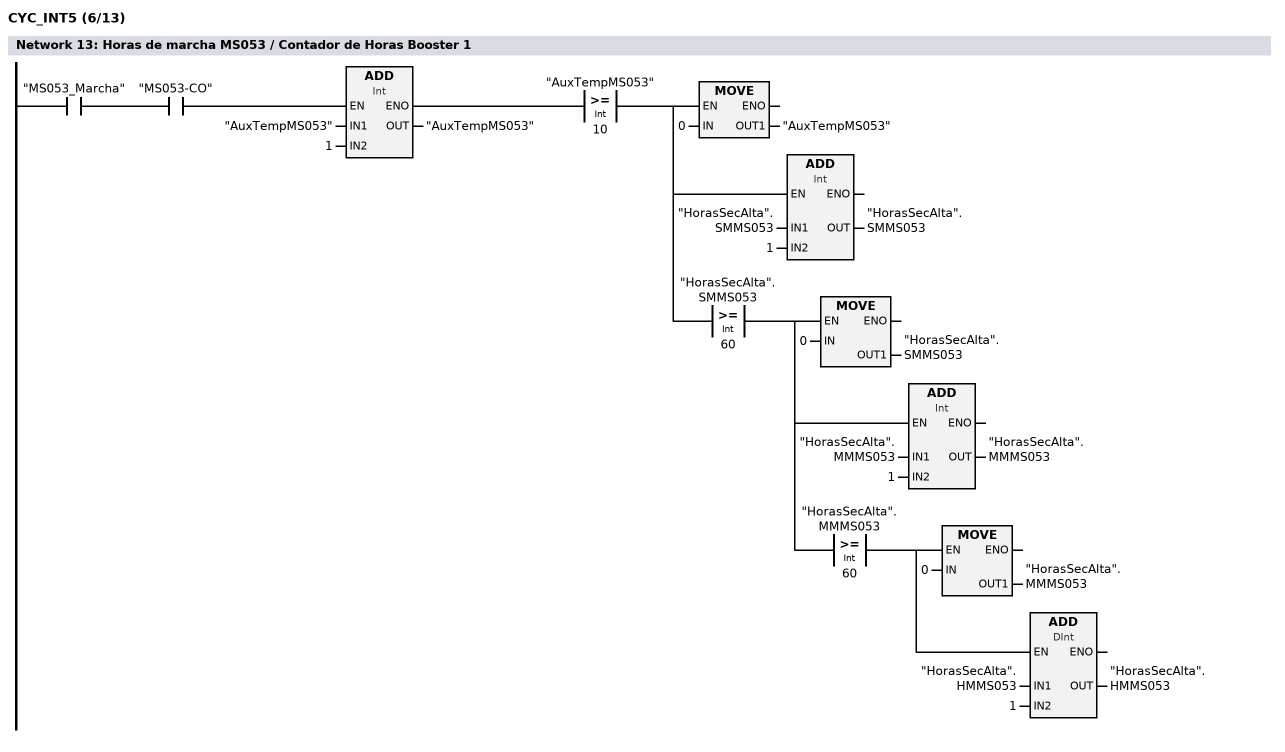
   RUNG wire#powerrail
      Contact( "MS053_Marcha" )
      Contact( "MS053-CO" )
      { S7_Templates := "SrcType := Int"; S7_GenerateENO := "TRUE" } Add(in1 := "AuxTempMS053", in2 := 1, out => "AuxTempMS053")
      { S7_Templates := "SrcType := Int" } GE_Contact(in1 := "AuxTempMS053", in2 := 10)
      wire#w1
      { S7_GenerateENO := "TRUE" } Move(in := 0, out1 => "AuxTempMS053")
   END_RUNG
   RUNG wire#w1
      { S7_Templates := "SrcType := Int"; S7_GenerateENO := "TRUE" } Add(in1 := "HorasSecAlta".SMMS053, in2 := 1, out => "HorasSecAlta".SMMS053)
   END_RUNG
   RUNG wire#w1
      { S7_Templates := "SrcType := Int" } GE_Contact(in1 := "HorasSecAlta".SMMS053, in2 := 60)
      wire#w2
      { S7_GenerateENO := "TRUE" } Move(in := 0, out1 => "HorasSecAlta".SMMS053)
   END_RUNG
   RUNG wire#w2
      { S7_Templates := "SrcType := Int"; S7_GenerateENO := "TRUE" } Add(in1 := "HorasSecAlta".MMMS053, in2 := 1, out => "HorasSecAlta".MMMS053)
   END_RUNG
   RUNG wire#w2
      { S7_Templates := "SrcType := Int" } GE_Contact(in1 := "HorasSecAlta".MMMS053, in2 := 60)
      wire#w3
      { S7_GenerateENO := "TRUE" } Move(in := 0, out1 => "HorasSecAlta".MMMS053)
   END_RUNG
   RUNG wire#w3
      { S7_Templates := "SrcType := DInt"; S7_GenerateENO := "TRUE" } Add(in1 := "HorasSecAlta".HMMS053, in2 := 1, out => "HorasSecAlta".HMMS053)
   END_RUNG
   // the same network as SCL:
   // ENO of a box is taken as its EN; it also drops when the box reports an error
   #_w1 := "MS053_Marcha" AND "MS053-CO";
   IF #_w1 THEN "AuxTempMS053" := "AuxTempMS053" + 1; END_IF;
   #_w2 := #_w1 AND ("AuxTempMS053" >= 10);
   IF #_w2 THEN
       "AuxTempMS053" := 0;
       "HorasSecAlta".SMMS053 := "HorasSecAlta".SMMS053 + 1;
   END_IF;
   #_w3 := #_w2 AND ("HorasSecAlta".SMMS053 >= 60);
   IF #_w3 THEN
       "HorasSecAlta".SMMS053 := 0;
       "HorasSecAlta".MMMS053 := "HorasSecAlta".MMMS053 + 1;
   END_IF;
   #_w4 := #_w3 AND ("HorasSecAlta".MMMS053 >= 60);
   IF #_w4 THEN
       "HorasSecAlta".MMMS053 := 0;
       "HorasSecAlta".HMMS053 := "HorasSecAlta".HMMS053 + 1;
   END_IF;
END_REGION

REGION Network 14: Horas de marcha MS054 / Contador de Horas Booster 1
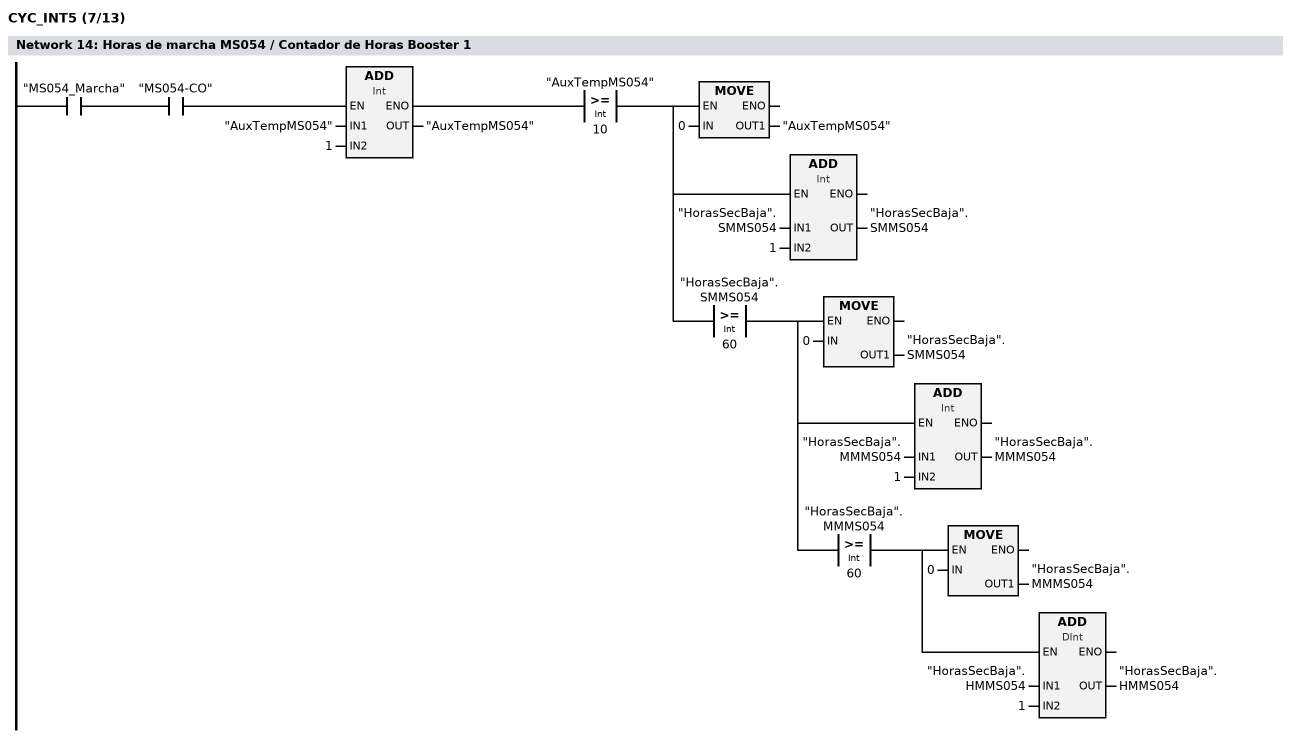
   RUNG wire#powerrail
      Contact( "MS054_Marcha" )
      Contact( "MS054-CO" )
      { S7_Templates := "SrcType := Int"; S7_GenerateENO := "TRUE" } Add(in1 := "AuxTempMS054", in2 := 1, out => "AuxTempMS054")
      { S7_Templates := "SrcType := Int" } GE_Contact(in1 := "AuxTempMS054", in2 := 10)
      wire#w1
      { S7_GenerateENO := "TRUE" } Move(in := 0, out1 => "AuxTempMS054")
   END_RUNG
   RUNG wire#w1
      { S7_Templates := "SrcType := Int"; S7_GenerateENO := "TRUE" } Add(in1 := "HorasSecBaja".SMMS054, in2 := 1, out => "HorasSecBaja".SMMS054)
   END_RUNG
   RUNG wire#w1
      { S7_Templates := "SrcType := Int" } GE_Contact(in1 := "HorasSecBaja".SMMS054, in2 := 60)
      wire#w2
      { S7_GenerateENO := "TRUE" } Move(in := 0, out1 => "HorasSecBaja".SMMS054)
   END_RUNG
   RUNG wire#w2
      { S7_Templates := "SrcType := Int"; S7_GenerateENO := "TRUE" } Add(in1 := "HorasSecBaja".MMMS054, in2 := 1, out => "HorasSecBaja".MMMS054)
   END_RUNG
   RUNG wire#w2
      { S7_Templates := "SrcType := Int" } GE_Contact(in1 := "HorasSecBaja".MMMS054, in2 := 60)
      wire#w3
      { S7_GenerateENO := "TRUE" } Move(in := 0, out1 => "HorasSecBaja".MMMS054)
   END_RUNG
   RUNG wire#w3
      { S7_Templates := "SrcType := DInt"; S7_GenerateENO := "TRUE" } Add(in1 := "HorasSecBaja".HMMS054, in2 := 1, out => "HorasSecBaja".HMMS054)
   END_RUNG
   // the same network as SCL:
   // ENO of a box is taken as its EN; it also drops when the box reports an error
   #_w1 := "MS054_Marcha" AND "MS054-CO";
   IF #_w1 THEN "AuxTempMS054" := "AuxTempMS054" + 1; END_IF;
   #_w2 := #_w1 AND ("AuxTempMS054" >= 10);
   IF #_w2 THEN
       "AuxTempMS054" := 0;
       "HorasSecBaja".SMMS054 := "HorasSecBaja".SMMS054 + 1;
   END_IF;
   #_w3 := #_w2 AND ("HorasSecBaja".SMMS054 >= 60);
   IF #_w3 THEN
       "HorasSecBaja".SMMS054 := 0;
       "HorasSecBaja".MMMS054 := "HorasSecBaja".MMMS054 + 1;
   END_IF;
   #_w4 := #_w3 AND ("HorasSecBaja".MMMS054 >= 60);
   IF #_w4 THEN
       "HorasSecBaja".MMMS054 := 0;
       "HorasSecBaja".HMMS054 := "HorasSecBaja".HMMS054 + 1;
   END_IF;
END_REGION

REGION Network 15: Horas de marcha MS055 / Contador de Horas Booster 1
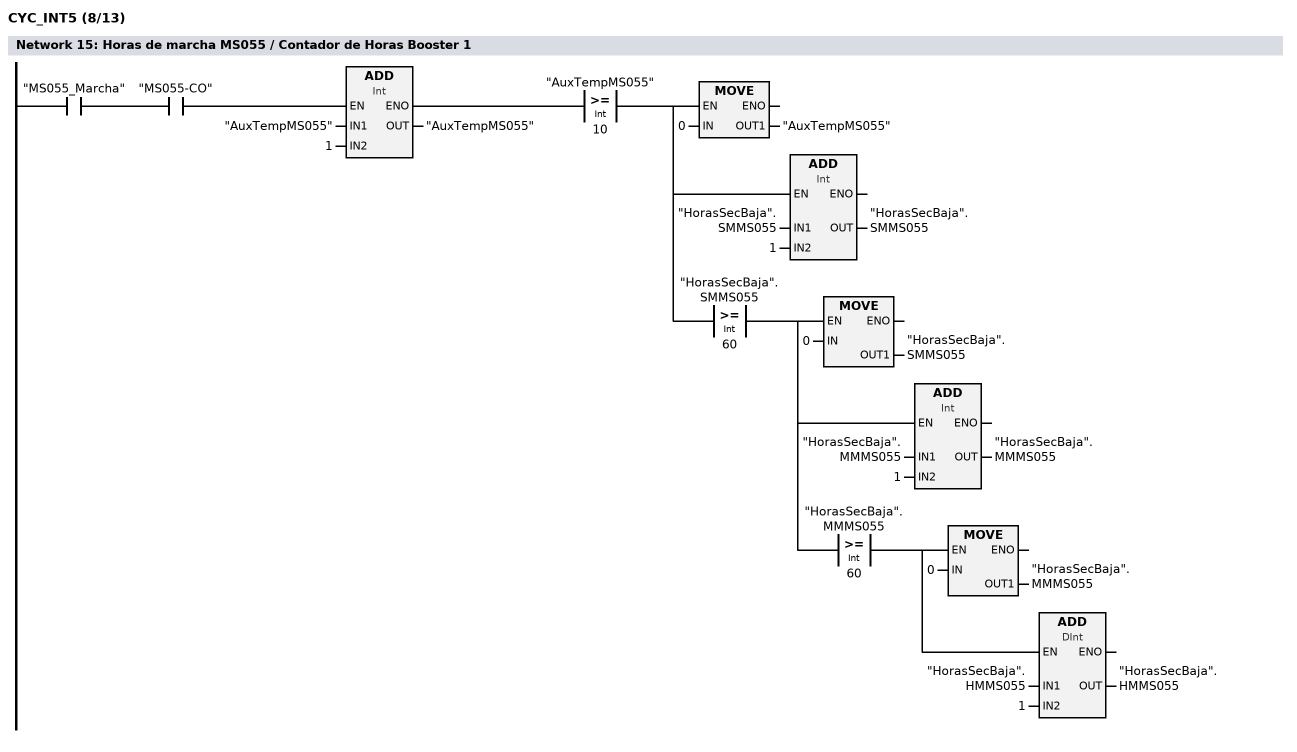
   RUNG wire#powerrail
      Contact( "MS055_Marcha" )
      Contact( "MS055-CO" )
      { S7_Templates := "SrcType := Int"; S7_GenerateENO := "TRUE" } Add(in1 := "AuxTempMS055", in2 := 1, out => "AuxTempMS055")
      { S7_Templates := "SrcType := Int" } GE_Contact(in1 := "AuxTempMS055", in2 := 10)
      wire#w1
      { S7_GenerateENO := "TRUE" } Move(in := 0, out1 => "AuxTempMS055")
   END_RUNG
   RUNG wire#w1
      { S7_Templates := "SrcType := Int"; S7_GenerateENO := "TRUE" } Add(in1 := "HorasSecBaja".SMMS055, in2 := 1, out => "HorasSecBaja".SMMS055)
   END_RUNG
   RUNG wire#w1
      { S7_Templates := "SrcType := Int" } GE_Contact(in1 := "HorasSecBaja".SMMS055, in2 := 60)
      wire#w2
      { S7_GenerateENO := "TRUE" } Move(in := 0, out1 => "HorasSecBaja".SMMS055)
   END_RUNG
   RUNG wire#w2
      { S7_Templates := "SrcType := Int"; S7_GenerateENO := "TRUE" } Add(in1 := "HorasSecBaja".MMMS055, in2 := 1, out => "HorasSecBaja".MMMS055)
   END_RUNG
   RUNG wire#w2
      { S7_Templates := "SrcType := Int" } GE_Contact(in1 := "HorasSecBaja".MMMS055, in2 := 60)
      wire#w3
      { S7_GenerateENO := "TRUE" } Move(in := 0, out1 => "HorasSecBaja".MMMS055)
   END_RUNG
   RUNG wire#w3
      { S7_Templates := "SrcType := DInt"; S7_GenerateENO := "TRUE" } Add(in1 := "HorasSecBaja".HMMS055, in2 := 1, out => "HorasSecBaja".HMMS055)
   END_RUNG
   // the same network as SCL:
   // ENO of a box is taken as its EN; it also drops when the box reports an error
   #_w1 := "MS055_Marcha" AND "MS055-CO";
   IF #_w1 THEN "AuxTempMS055" := "AuxTempMS055" + 1; END_IF;
   #_w2 := #_w1 AND ("AuxTempMS055" >= 10);
   IF #_w2 THEN
       "AuxTempMS055" := 0;
       "HorasSecBaja".SMMS055 := "HorasSecBaja".SMMS055 + 1;
   END_IF;
   #_w3 := #_w2 AND ("HorasSecBaja".SMMS055 >= 60);
   IF #_w3 THEN
       "HorasSecBaja".SMMS055 := 0;
       "HorasSecBaja".MMMS055 := "HorasSecBaja".MMMS055 + 1;
   END_IF;
   #_w4 := #_w3 AND ("HorasSecBaja".MMMS055 >= 60);
   IF #_w4 THEN
       "HorasSecBaja".MMMS055 := 0;
       "HorasSecBaja".HMMS055 := "HorasSecBaja".HMMS055 + 1;
   END_IF;
END_REGION

REGION Network 16: Horas de marcha MC060 / Contador de Horas Booster 1
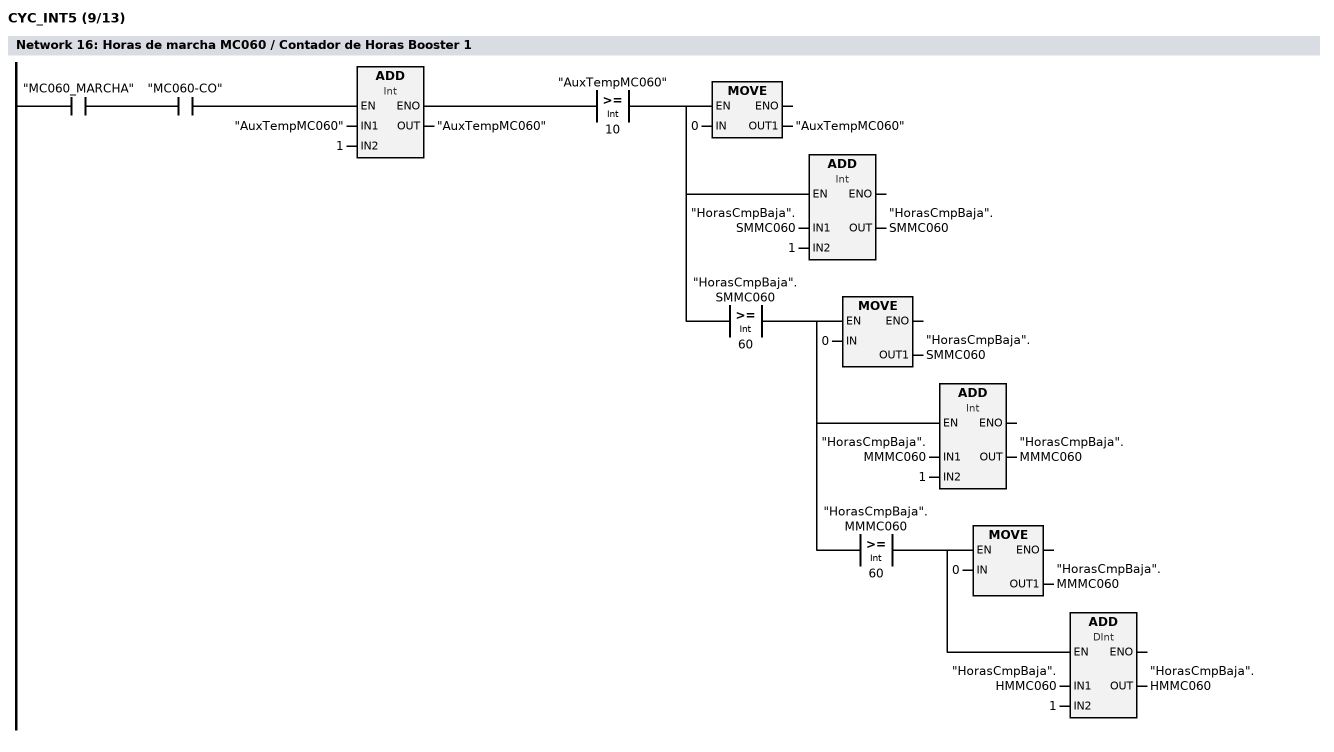
   RUNG wire#powerrail
      Contact( "MC060_MARCHA" )
      Contact( "MC060-CO" )
      { S7_Templates := "SrcType := Int"; S7_GenerateENO := "TRUE" } Add(in1 := "AuxTempMC060", in2 := 1, out => "AuxTempMC060")
      { S7_Templates := "SrcType := Int" } GE_Contact(in1 := "AuxTempMC060", in2 := 10)
      wire#w1
      { S7_GenerateENO := "TRUE" } Move(in := 0, out1 => "AuxTempMC060")
   END_RUNG
   RUNG wire#w1
      { S7_Templates := "SrcType := Int"; S7_GenerateENO := "TRUE" } Add(in1 := "HorasCmpBaja".SMMC060, in2 := 1, out => "HorasCmpBaja".SMMC060)
   END_RUNG
   RUNG wire#w1
      { S7_Templates := "SrcType := Int" } GE_Contact(in1 := "HorasCmpBaja".SMMC060, in2 := 60)
      wire#w2
      { S7_GenerateENO := "TRUE" } Move(in := 0, out1 => "HorasCmpBaja".SMMC060)
   END_RUNG
   RUNG wire#w2
      { S7_Templates := "SrcType := Int"; S7_GenerateENO := "TRUE" } Add(in1 := "HorasCmpBaja".MMMC060, in2 := 1, out => "HorasCmpBaja".MMMC060)
   END_RUNG
   RUNG wire#w2
      { S7_Templates := "SrcType := Int" } GE_Contact(in1 := "HorasCmpBaja".MMMC060, in2 := 60)
      wire#w3
      { S7_GenerateENO := "TRUE" } Move(in := 0, out1 => "HorasCmpBaja".MMMC060)
   END_RUNG
   RUNG wire#w3
      { S7_Templates := "SrcType := DInt"; S7_GenerateENO := "TRUE" } Add(in1 := "HorasCmpBaja".HMMC060, in2 := 1, out => "HorasCmpBaja".HMMC060)
   END_RUNG
   // the same network as SCL:
   // ENO of a box is taken as its EN; it also drops when the box reports an error
   #_w1 := "MC060_MARCHA" AND "MC060-CO";
   IF #_w1 THEN "AuxTempMC060" := "AuxTempMC060" + 1; END_IF;
   #_w2 := #_w1 AND ("AuxTempMC060" >= 10);
   IF #_w2 THEN
       "AuxTempMC060" := 0;
       "HorasCmpBaja".SMMC060 := "HorasCmpBaja".SMMC060 + 1;
   END_IF;
   #_w3 := #_w2 AND ("HorasCmpBaja".SMMC060 >= 60);
   IF #_w3 THEN
       "HorasCmpBaja".SMMC060 := 0;
       "HorasCmpBaja".MMMC060 := "HorasCmpBaja".MMMC060 + 1;
   END_IF;
   #_w4 := #_w3 AND ("HorasCmpBaja".MMMC060 >= 60);
   IF #_w4 THEN
       "HorasCmpBaja".MMMC060 := 0;
       "HorasCmpBaja".HMMC060 := "HorasCmpBaja".HMMC060 + 1;
   END_IF;
END_REGION

REGION Network 17: Horas de marcha MC061 / Contador de Horas Booster 1
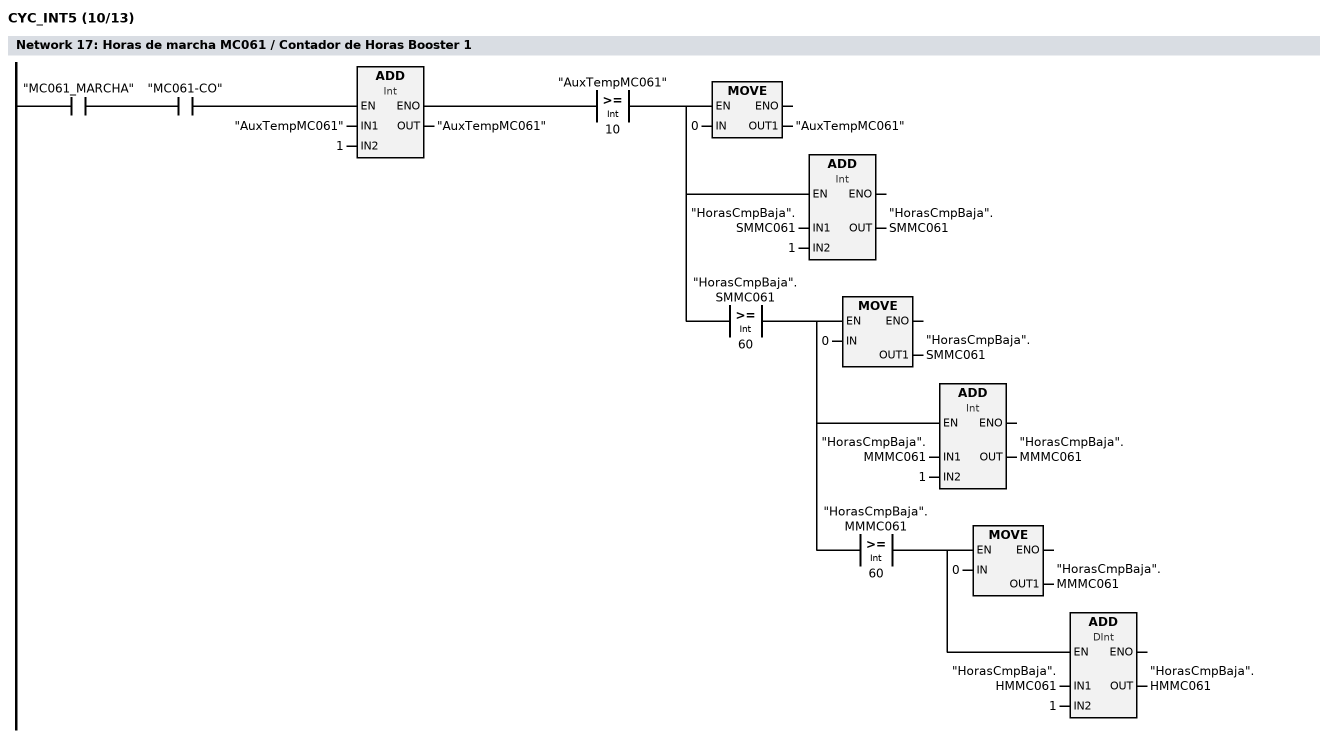
   RUNG wire#powerrail
      Contact( "MC061_MARCHA" )
      Contact( "MC061-CO" )
      { S7_Templates := "SrcType := Int"; S7_GenerateENO := "TRUE" } Add(in1 := "AuxTempMC061", in2 := 1, out => "AuxTempMC061")
      { S7_Templates := "SrcType := Int" } GE_Contact(in1 := "AuxTempMC061", in2 := 10)
      wire#w1
      { S7_GenerateENO := "TRUE" } Move(in := 0, out1 => "AuxTempMC061")
   END_RUNG
   RUNG wire#w1
      { S7_Templates := "SrcType := Int"; S7_GenerateENO := "TRUE" } Add(in1 := "HorasCmpBaja".SMMC061, in2 := 1, out => "HorasCmpBaja".SMMC061)
   END_RUNG
   RUNG wire#w1
      { S7_Templates := "SrcType := Int" } GE_Contact(in1 := "HorasCmpBaja".SMMC061, in2 := 60)
      wire#w2
      { S7_GenerateENO := "TRUE" } Move(in := 0, out1 => "HorasCmpBaja".SMMC061)
   END_RUNG
   RUNG wire#w2
      { S7_Templates := "SrcType := Int"; S7_GenerateENO := "TRUE" } Add(in1 := "HorasCmpBaja".MMMC061, in2 := 1, out => "HorasCmpBaja".MMMC061)
   END_RUNG
   RUNG wire#w2
      { S7_Templates := "SrcType := Int" } GE_Contact(in1 := "HorasCmpBaja".MMMC061, in2 := 60)
      wire#w3
      { S7_GenerateENO := "TRUE" } Move(in := 0, out1 => "HorasCmpBaja".MMMC061)
   END_RUNG
   RUNG wire#w3
      { S7_Templates := "SrcType := DInt"; S7_GenerateENO := "TRUE" } Add(in1 := "HorasCmpBaja".HMMC061, in2 := 1, out => "HorasCmpBaja".HMMC061)
   END_RUNG
   // the same network as SCL:
   // ENO of a box is taken as its EN; it also drops when the box reports an error
   #_w1 := "MC061_MARCHA" AND "MC061-CO";
   IF #_w1 THEN "AuxTempMC061" := "AuxTempMC061" + 1; END_IF;
   #_w2 := #_w1 AND ("AuxTempMC061" >= 10);
   IF #_w2 THEN
       "AuxTempMC061" := 0;
       "HorasCmpBaja".SMMC061 := "HorasCmpBaja".SMMC061 + 1;
   END_IF;
   #_w3 := #_w2 AND ("HorasCmpBaja".SMMC061 >= 60);
   IF #_w3 THEN
       "HorasCmpBaja".SMMC061 := 0;
       "HorasCmpBaja".MMMC061 := "HorasCmpBaja".MMMC061 + 1;
   END_IF;
   #_w4 := #_w3 AND ("HorasCmpBaja".MMMC061 >= 60);
   IF #_w4 THEN
       "HorasCmpBaja".MMMC061 := 0;
       "HorasCmpBaja".HMMC061 := "HorasCmpBaja".HMMC061 + 1;
   END_IF;
END_REGION

REGION Network 18: Horas de marcha MC062 / Contador de Horas Booster 1
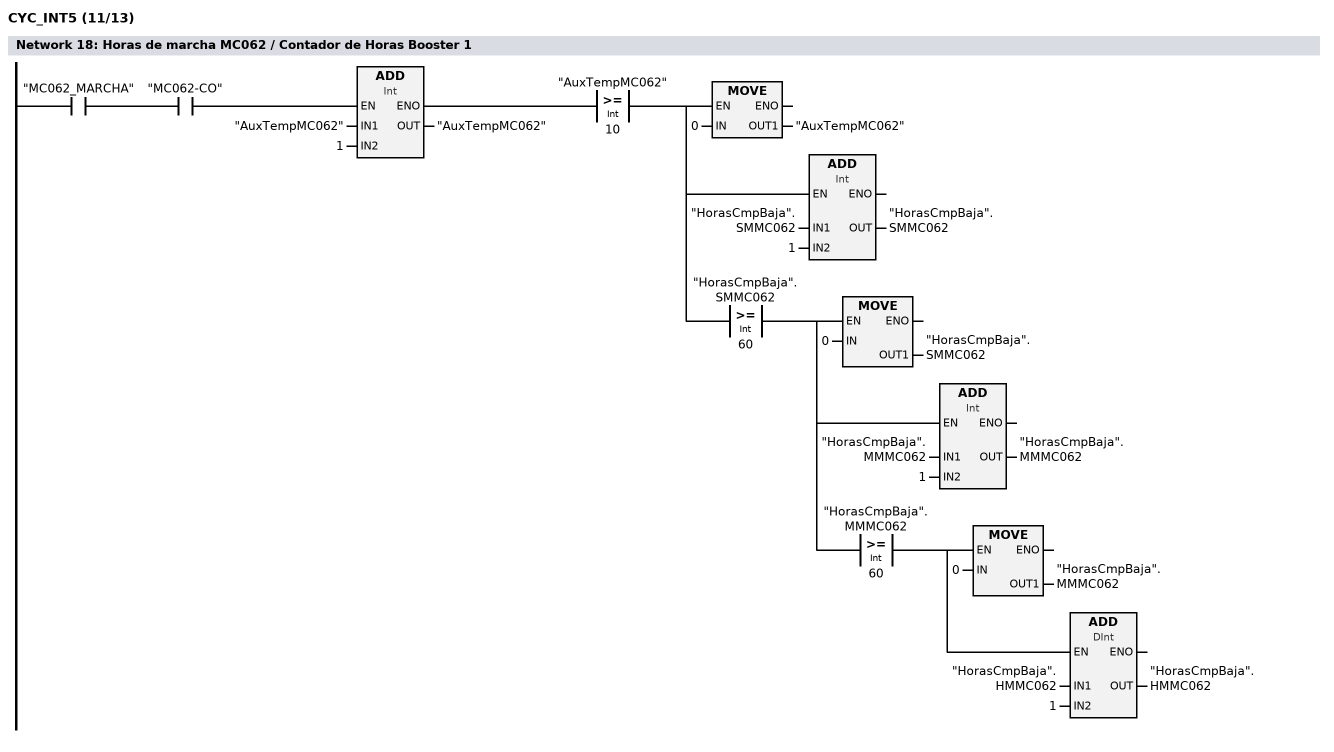
   RUNG wire#powerrail
      Contact( "MC062_MARCHA" )
      Contact( "MC062-CO" )
      { S7_Templates := "SrcType := Int"; S7_GenerateENO := "TRUE" } Add(in1 := "AuxTempMC062", in2 := 1, out => "AuxTempMC062")
      { S7_Templates := "SrcType := Int" } GE_Contact(in1 := "AuxTempMC062", in2 := 10)
      wire#w1
      { S7_GenerateENO := "TRUE" } Move(in := 0, out1 => "AuxTempMC062")
   END_RUNG
   RUNG wire#w1
      { S7_Templates := "SrcType := Int"; S7_GenerateENO := "TRUE" } Add(in1 := "HorasCmpBaja".SMMC062, in2 := 1, out => "HorasCmpBaja".SMMC062)
   END_RUNG
   RUNG wire#w1
      { S7_Templates := "SrcType := Int" } GE_Contact(in1 := "HorasCmpBaja".SMMC062, in2 := 60)
      wire#w2
      { S7_GenerateENO := "TRUE" } Move(in := 0, out1 => "HorasCmpBaja".SMMC062)
   END_RUNG
   RUNG wire#w2
      { S7_Templates := "SrcType := Int"; S7_GenerateENO := "TRUE" } Add(in1 := "HorasCmpBaja".MMMC062, in2 := 1, out => "HorasCmpBaja".MMMC062)
   END_RUNG
   RUNG wire#w2
      { S7_Templates := "SrcType := Int" } GE_Contact(in1 := "HorasCmpBaja".MMMC062, in2 := 60)
      wire#w3
      { S7_GenerateENO := "TRUE" } Move(in := 0, out1 => "HorasCmpBaja".MMMC062)
   END_RUNG
   RUNG wire#w3
      { S7_Templates := "SrcType := DInt"; S7_GenerateENO := "TRUE" } Add(in1 := "HorasCmpBaja".HMMC062, in2 := 1, out => "HorasCmpBaja".HMMC062)
   END_RUNG
   // the same network as SCL:
   // ENO of a box is taken as its EN; it also drops when the box reports an error
   #_w1 := "MC062_MARCHA" AND "MC062-CO";
   IF #_w1 THEN "AuxTempMC062" := "AuxTempMC062" + 1; END_IF;
   #_w2 := #_w1 AND ("AuxTempMC062" >= 10);
   IF #_w2 THEN
       "AuxTempMC062" := 0;
       "HorasCmpBaja".SMMC062 := "HorasCmpBaja".SMMC062 + 1;
   END_IF;
   #_w3 := #_w2 AND ("HorasCmpBaja".SMMC062 >= 60);
   IF #_w3 THEN
       "HorasCmpBaja".SMMC062 := 0;
       "HorasCmpBaja".MMMC062 := "HorasCmpBaja".MMMC062 + 1;
   END_IF;
   #_w4 := #_w3 AND ("HorasCmpBaja".MMMC062 >= 60);
   IF #_w4 THEN
       "HorasCmpBaja".MMMC062 := 0;
       "HorasCmpBaja".HMMC062 := "HorasCmpBaja".HMMC062 + 1;
   END_IF;
END_REGION

REGION Network 19: Horas de marcha MC063 / Contador de Horas Booster 1
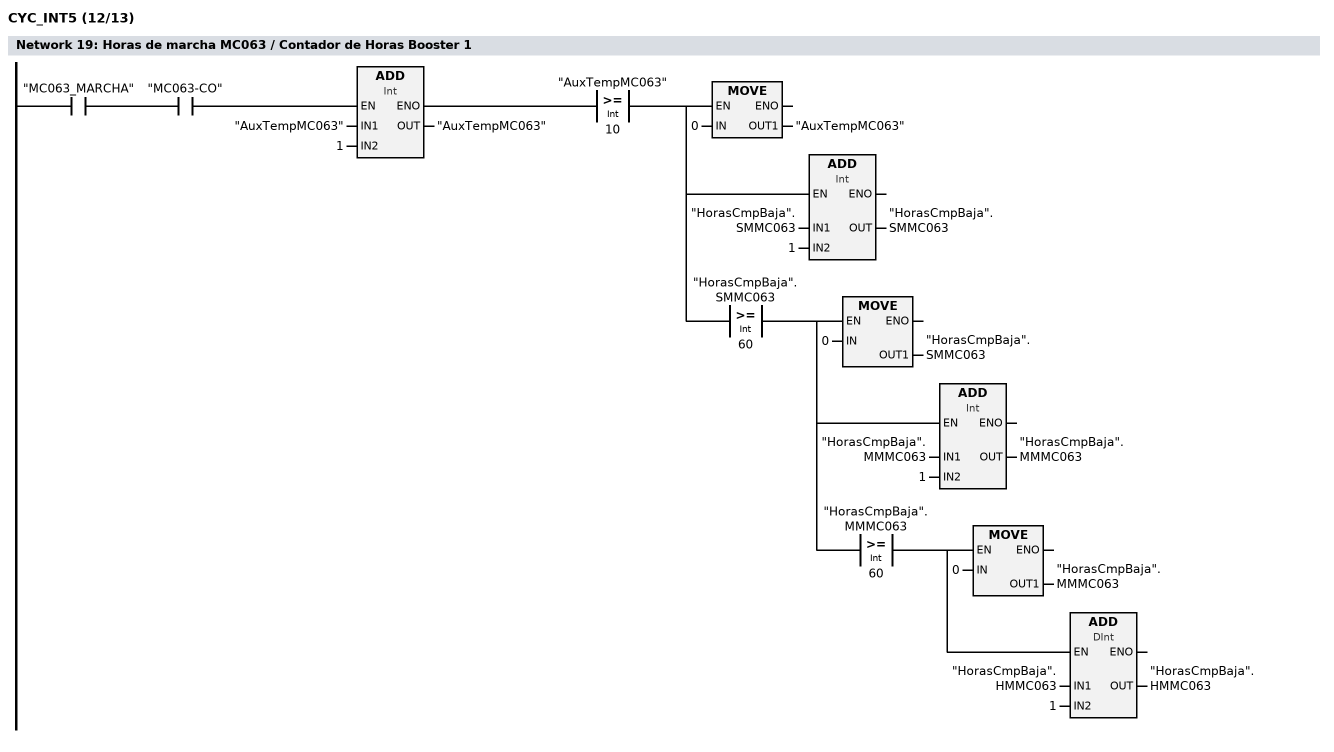
   RUNG wire#powerrail
      Contact( "MC063_MARCHA" )
      Contact( "MC063-CO" )
      { S7_Templates := "SrcType := Int"; S7_GenerateENO := "TRUE" } Add(in1 := "AuxTempMC063", in2 := 1, out => "AuxTempMC063")
      { S7_Templates := "SrcType := Int" } GE_Contact(in1 := "AuxTempMC063", in2 := 10)
      wire#w1
      { S7_GenerateENO := "TRUE" } Move(in := 0, out1 => "AuxTempMC063")
   END_RUNG
   RUNG wire#w1
      { S7_Templates := "SrcType := Int"; S7_GenerateENO := "TRUE" } Add(in1 := "HorasCmpBaja".SMMC063, in2 := 1, out => "HorasCmpBaja".SMMC063)
   END_RUNG
   RUNG wire#w1
      { S7_Templates := "SrcType := Int" } GE_Contact(in1 := "HorasCmpBaja".SMMC063, in2 := 60)
      wire#w2
      { S7_GenerateENO := "TRUE" } Move(in := 0, out1 => "HorasCmpBaja".SMMC063)
   END_RUNG
   RUNG wire#w2
      { S7_Templates := "SrcType := Int"; S7_GenerateENO := "TRUE" } Add(in1 := "HorasCmpBaja".MMMC063, in2 := 1, out => "HorasCmpBaja".MMMC063)
   END_RUNG
   RUNG wire#w2
      { S7_Templates := "SrcType := Int" } GE_Contact(in1 := "HorasCmpBaja".MMMC063, in2 := 60)
      wire#w3
      { S7_GenerateENO := "TRUE" } Move(in := 0, out1 => "HorasCmpBaja".MMMC063)
   END_RUNG
   RUNG wire#w3
      { S7_Templates := "SrcType := DInt"; S7_GenerateENO := "TRUE" } Add(in1 := "HorasCmpBaja".HMMC063, in2 := 1, out => "HorasCmpBaja".HMMC063)
   END_RUNG
   // the same network as SCL:
   // ENO of a box is taken as its EN; it also drops when the box reports an error
   #_w1 := "MC063_MARCHA" AND "MC063-CO";
   IF #_w1 THEN "AuxTempMC063" := "AuxTempMC063" + 1; END_IF;
   #_w2 := #_w1 AND ("AuxTempMC063" >= 10);
   IF #_w2 THEN
       "AuxTempMC063" := 0;
       "HorasCmpBaja".SMMC063 := "HorasCmpBaja".SMMC063 + 1;
   END_IF;
   #_w3 := #_w2 AND ("HorasCmpBaja".SMMC063 >= 60);
   IF #_w3 THEN
       "HorasCmpBaja".SMMC063 := 0;
       "HorasCmpBaja".MMMC063 := "HorasCmpBaja".MMMC063 + 1;
   END_IF;
   #_w4 := #_w3 AND ("HorasCmpBaja".MMMC063 >= 60);
   IF #_w4 THEN
       "HorasCmpBaja".MMMC063 := 0;
       "HorasCmpBaja".HMMC063 := "HorasCmpBaja".HMMC063 + 1;
   END_IF;
END_REGION

REGION Network 20: Horas de marcha MC064 / Contador de Horas Booster 1
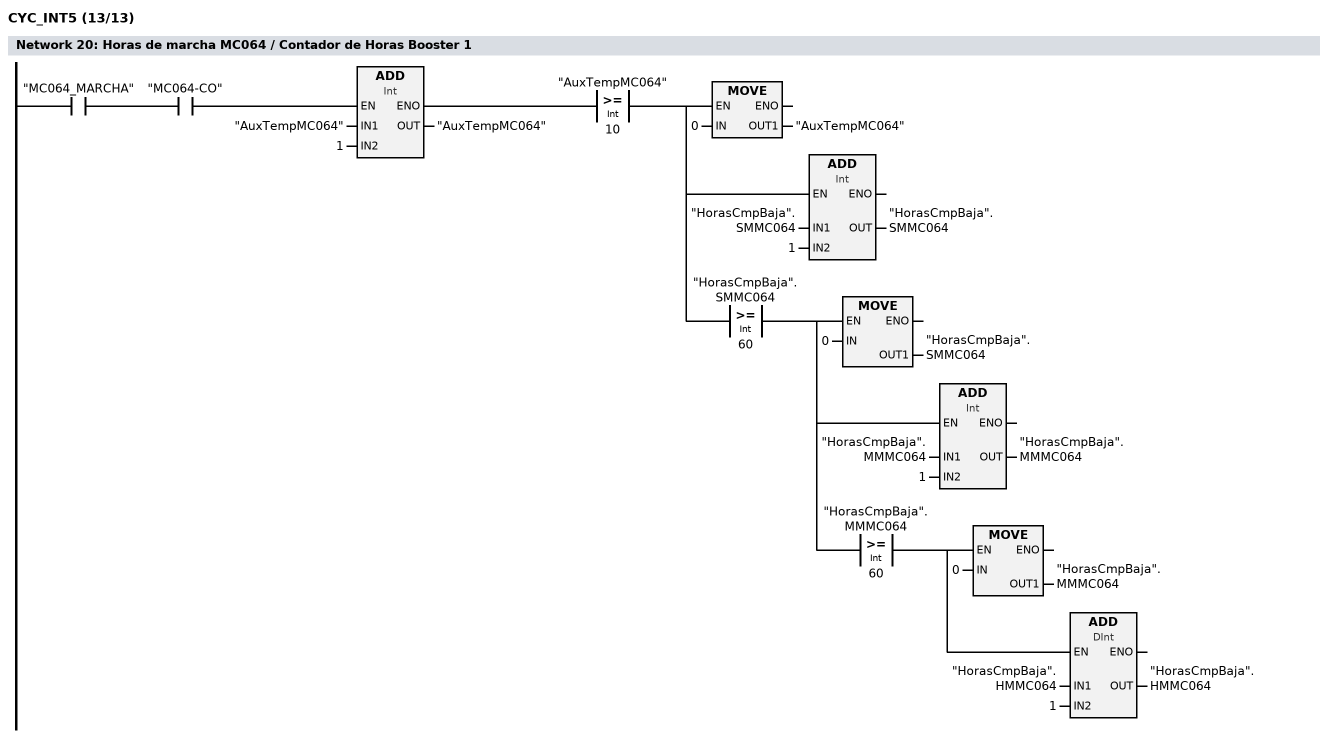
   RUNG wire#powerrail
      Contact( "MC064_MARCHA" )
      Contact( "MC064-CO" )
      { S7_Templates := "SrcType := Int"; S7_GenerateENO := "TRUE" } Add(in1 := "AuxTempMC064", in2 := 1, out => "AuxTempMC064")
      { S7_Templates := "SrcType := Int" } GE_Contact(in1 := "AuxTempMC064", in2 := 10)
      wire#w1
      { S7_GenerateENO := "TRUE" } Move(in := 0, out1 => "AuxTempMC064")
   END_RUNG
   RUNG wire#w1
      { S7_Templates := "SrcType := Int"; S7_GenerateENO := "TRUE" } Add(in1 := "HorasCmpBaja".SMMC064, in2 := 1, out => "HorasCmpBaja".SMMC064)
   END_RUNG
   RUNG wire#w1
      { S7_Templates := "SrcType := Int" } GE_Contact(in1 := "HorasCmpBaja".SMMC064, in2 := 60)
      wire#w2
      { S7_GenerateENO := "TRUE" } Move(in := 0, out1 => "HorasCmpBaja".SMMC064)
   END_RUNG
   RUNG wire#w2
      { S7_Templates := "SrcType := Int"; S7_GenerateENO := "TRUE" } Add(in1 := "HorasCmpBaja".MMMC064, in2 := 1, out => "HorasCmpBaja".MMMC064)
   END_RUNG
   RUNG wire#w2
      { S7_Templates := "SrcType := Int" } GE_Contact(in1 := "HorasCmpBaja".MMMC064, in2 := 60)
      wire#w3
      { S7_GenerateENO := "TRUE" } Move(in := 0, out1 => "HorasCmpBaja".MMMC064)
   END_RUNG
   RUNG wire#w3
      { S7_Templates := "SrcType := DInt"; S7_GenerateENO := "TRUE" } Add(in1 := "HorasCmpBaja".HMMC064, in2 := 1, out => "HorasCmpBaja".HMMC064)
   END_RUNG
   // the same network as SCL:
   // ENO of a box is taken as its EN; it also drops when the box reports an error
   #_w1 := "MC064_MARCHA" AND "MC064-CO";
   IF #_w1 THEN "AuxTempMC064" := "AuxTempMC064" + 1; END_IF;
   #_w2 := #_w1 AND ("AuxTempMC064" >= 10);
   IF #_w2 THEN
       "AuxTempMC064" := 0;
       "HorasCmpBaja".SMMC064 := "HorasCmpBaja".SMMC064 + 1;
   END_IF;
   #_w3 := #_w2 AND ("HorasCmpBaja".SMMC064 >= 60);
   IF #_w3 THEN
       "HorasCmpBaja".SMMC064 := 0;
       "HorasCmpBaja".MMMC064 := "HorasCmpBaja".MMMC064 + 1;
   END_IF;
   #_w4 := #_w3 AND ("HorasCmpBaja".MMMC064 >= 60);
   IF #_w4 THEN
       "HorasCmpBaja".MMMC064 := 0;
       "HorasCmpBaja".HMMC064 := "HorasCmpBaja".HMMC064 + 1;
   END_IF;
END_REGION
END_ORGANIZATION_BLOCK

// folder: Iluminación

FUNCTION "IluminaciónMTA" : Void   // FC23, LAD
{ S7_Optimized_Access := 'FALSE' }
VERSION : 0.1
   VAR_TEMP   // added for the SCL form of the ladder/FBD networks
      _s5time1 : S5Time;
      _w1 : Bool;
   END_VAR
BEGIN

REGION Network 1
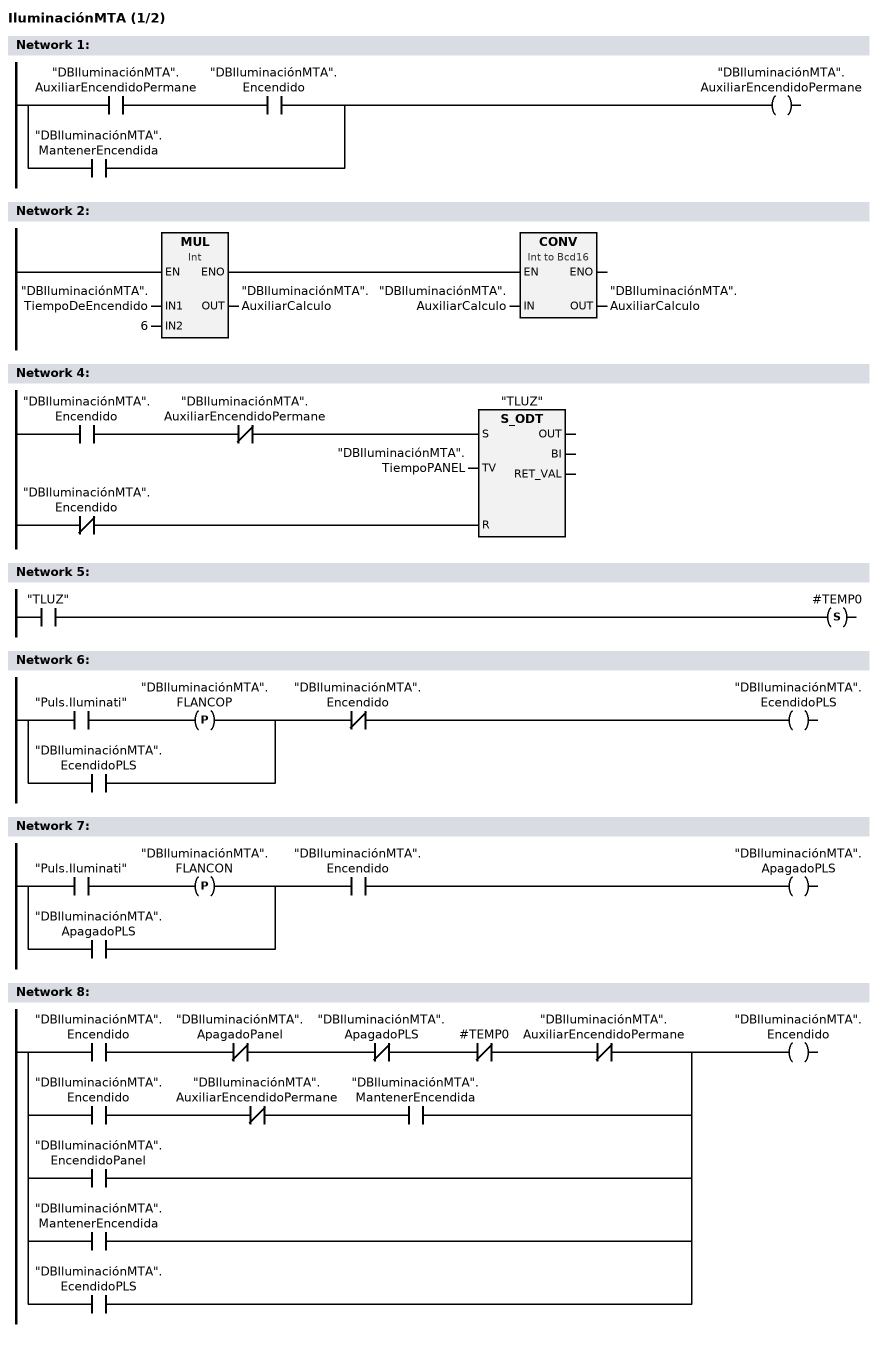
   "DBIluminaciónMTA".AuxiliarEncendidoPermane := "DBIluminaciónMTA".MantenerEncendida OR ("DBIluminaciónMTA".AuxiliarEncendidoPermane AND "DBIluminaciónMTA".Encendido);
END_REGION

REGION Network 2
   RUNG wire#powerrail
      { S7_Templates := "SrcType := Int"; S7_GenerateENO := "TRUE" } Mul(in1 := "DBIluminaciónMTA".TiempoDeEncendido, in2 := 6, out => "DBIluminaciónMTA".AuxiliarCalculo)
      { S7_Templates := "[SrcType := Int, DestType := Bcd16]"; S7_GenerateENO := "TRUE" } Convert(in := "DBIluminaciónMTA".AuxiliarCalculo, out => "DBIluminaciónMTA".AuxiliarCalculo)
   END_RUNG
   // the same network as SCL:
   // ENO of a box is taken as its EN; it also drops when the box reports an error
   "DBIluminaciónMTA".AuxiliarCalculo := "DBIluminaciónMTA".TiempoDeEncendido * 6;
   "DBIluminaciónMTA".AuxiliarCalculo := INT_TO_BCD16("DBIluminaciónMTA".AuxiliarCalculo);
END_REGION
